
screen "Dev_VD2" 800x480, template "Settings"
   TextField "Text field_10" at 472,32 size 34x18; Text 'ОС.О'
   TextField "Text field_4" at 510,10 size 77x22; Text 'Сигналы:'
   Button "Button_21" at 508,32 size 60x20; TextOff 'Text'; Authorization "User administration"; PictureList "ON_OFF"
      on Click: InvertBit("V_x_Use_Open")
      ProcessValue <- "V_x_Use_Open"
   Button "Button_22" at 508,56 size 60x20; TextOff 'Text'; PictureList "ON_OFF"; Authorization "User administration"
      on Click: InvertBit("V_x_Use_Close")
      ProcessValue <- "V_x_Use_Close"
   Button "Button_27" at 452,31 size 20x20; TextOff 'Text'; Authorization "User administration"; PictureList "signal_green"
      ProcessValue <- "V_x_FB_Open"
   GraphicIOField "Graphic I/O field_5" at 169,56 size 50x50; PictureList "Valve_Hor"
      ProcessValue <- "V_x_Status"
   TextField "Text field_6" at 472,56 size 31x18; Text 'ОС.З'
   Button "Button_12" at 452,55 size 20x20; TextOff 'Text'; Authorization "User administration"; PictureList "signal_green"
      ProcessValue <- "V_x_FB_Close"
   Button "Button_2" at 574,32 size 20x20; TextOff 'Text'; Authorization "User administration"; PictureList "ok_green"
      on Release: InvertBit("V_x_Inv_Open")
      ProcessValue <- "V_x_Inv_Open"
   Button "Button_3" at 574,56 size 20x20; TextOff 'Text'; Authorization "User administration"; PictureList "ok_green"
      on Release: InvertBit("V_x_Inv_Close")
      ProcessValue <- "V_x_Inv_Close"
   IOField "I/O field_1" at 615,30 size 30x24; Authorization "Developer"; FormatPattern 99
      ProcessValue <- "V_x_Indirect_BYTE_FB_Open"
   IOField "I/O field_6" at 655,30 size 20x24; Authorization "Developer"; FormatPattern 9
      ProcessValue <- "V_x_Indirect_BIT_FB_Open"
   TextField "Text field_11" at 601,30 size 13x23; Text 'I'
   TextField "Text field_1" at 644,30 size 13x23; Text '.'
   IOField "I/O field_2" at 615,54 size 30x24; Authorization "Developer"; FormatPattern 99
      ProcessValue <- "V_x_Indirect_BYTE_FB_Close"
   IOField "I/O field_3" at 655,54 size 20x24; Authorization "Developer"; FormatPattern 9
      ProcessValue <- "V_x_Indirect_BIT_FB_Close"
   TextField "Text field_7" at 601,54 size 13x23; Text 'I'
   TextField "Text field_8" at 644,54 size 13x23; Text '.'
   IOField "I/O field_4" at 615,78 size 30x24; Authorization "Developer"; FormatPattern 99
      ProcessValue <- "V_x_Indirect_BYTE_CMD_Open"
   IOField "I/O field_7" at 655,78 size 20x24; Authorization "Developer"; FormatPattern 9
      ProcessValue <- "V_x_Indirect_BIT_CMD_Open"
   TextField "Text field_9" at 599,78 size 17x23; Text 'Q'
   TextField "Text field_13" at 644,78 size 13x23; Text '.'
   TextField "Text field_3" at 472,80 size 65x18; Text 'Открыть / CMD Откр'
   Button "Button_5" at 452,79 size 20x20; TextOff 'Text'; Authorization "User administration"; PictureList "signal_green"
      ProcessValue <- "V_x_CMD_Open"
   IOField "I/O field_8" at 170,11 size 171x26; FormatPattern ????????????????
      ProcessValue <- "Vx_Name"
   Button "Button_14" at 538,142 size 142x20; TextOff 'Фиксация'; Authorization "User administration"; TextList "Air_V"
      on Click: InvertBit("V_x_Use_Electro")
      Appearance <- "V_x_Use_Electro"
      ProcessValue <- "V_x_Use_Electro"
   Button "Button_28" at 540,80 size 60x20; TextOff 'Text'; Authorization "User administration"; PictureList "ON_OFF"
      on Click: InvertBit("V_x_Use_CMD_Open")
      ProcessValue <- "V_x_Use_CMD_Open"
   IOField "I/O field_9" at 615,102 size 30x24; Authorization "Developer"; FormatPattern 99
      ProcessValue <- "V_x_Indirect_BYTE_CMD_Close"
   IOField "I/O field_10" at 655,102 size 20x24; Authorization "Developer"; FormatPattern 9
      ProcessValue <- "V_x_Indirect_BIT_CMD_Close"
   TextField "Text field_12" at 599,102 size 17x23; Text 'Q'
   TextField "Text field_14" at 644,102 size 13x23; Text '.'
   TextField "Text field_16" at 472,104 size 62x18; Text 'Закрыть / CMD Закр'
   Button "Button_20" at 452,103 size 20x20; TextOff 'Text'; Authorization "User administration"; PictureList "signal_green"
      ProcessValue <- "V_x_CMD_Close"
   Button "Button_30" at 539,108 size 60x20; TextOff 'Text'; PictureList "ON_OFF"; Authorization "User administration"
      on Click: InvertBit("V_x_Use_CMD_Close")
      ProcessValue <- "V_x_Use_CMD_Close"
   Button "Button_1" at 165,265 size 112x32; TextOff 'DB 700'; Authorization "User administration"
      on Release: SetTag("Vx", 700); SetTag("Vx_Name", 'DB 700')
      Visibility <- "Support_DB_All_VD2s"
      Appearance <- "Vx"
   Button "Button_4" at 165,305 size 112x32; TextOff 'DB 701'; Authorization "User administration"
      on Release: SetTag("Vx", 701); SetTag("Vx_Name", 'DB 701')
      Visibility <- "Support_DB_All_VD2s"
      Appearance <- "Vx"
   Button "Button_17" at 165,345 size 112x32; TextOff 'DB 702'; Authorization "User administration"
      on Release: SetTag("Vx", 702); SetTag("Vx_Name", 'DB 702')
      Visibility <- "Support_DB_All_VD2s"
      Appearance <- "Vx"
   Button "Button_6" at 165,385 size 112x32; TextOff 'DB 703'; Authorization "User administration"
      on Release: SetTag("Vx", 703); SetTag("Vx_Name", 'DB 703')
      Visibility <- "Support_DB_All_VD2s"
      Appearance <- "Vx"
   Button "Button_15" at 443,265 size 112x32; TextOff 'DB 710'; Authorization "User administration"
      on Release: SetTag("Vx", 710); SetTag("Vx_Name", 'DB 710')
      Visibility <- "Support_DB_All_VD2s"
      Appearance <- "Vx"
   Button "Button_18" at 443,305 size 112x32; TextOff 'DB 711'; Authorization "User administration"
      on Release: SetTag("Vx", 711); SetTag("Vx_Name", 'DB 711')
      Visibility <- "Support_DB_All_VD2s"
      Appearance <- "Vx"
   Button "Button_23" at 443,345 size 112x32; TextOff 'DB 712'; Authorization "User administration"
      on Release: SetTag("Vx", 712); SetTag("Vx_Name", 'DB 712')
      Visibility <- "Support_DB_All_VD2s"
      Appearance <- "Vx"
   Button "Button_24" at 443,385 size 112x32; TextOff 'DB 713'; Authorization "User administration"
      on Release: SetTag("Vx", 713); SetTag("Vx_Name", 'DB 713')
      Visibility <- "Support_DB_All_VD2s"
      Appearance <- "Vx"
   Button "Button_25" at 443,425 size 112x32; TextOff 'DB 714'; Authorization "User administration"
      on Release: SetTag("Vx", 714); SetTag("Vx_Name", 'DB 714')
      Visibility <- "Support_DB_All_VD2s"
      Appearance <- "Vx"
   Button "Button_26" at 583,344 size 112x32; TextOff 'DB 717'; Authorization "User administration"
      on Release: SetTag("Vx", 717); SetTag("Vx_Name", 'DB 717')
      Visibility <- "Support_DB_All_VD2s"
      Appearance <- "Vx"
   Button "Button_29" at 583,384 size 112x32; TextOff 'DB 718'; Authorization "User administration"
      on Release: SetTag("Vx", 718); SetTag("Vx_Name", 'DB 718')
      Visibility <- "Support_DB_All_VD2s"
      Appearance <- "Vx"
   Button "Button_31" at 583,264 size 112x32; TextOff 'DB 715'; Authorization "User administration"
      on Release: SetTag("Vx", 715); SetTag("Vx_Name", 'DB 715')
      Visibility <- "Support_DB_All_VD2s"
      Appearance <- "Vx"
   Button "Button_32" at 583,304 size 112x32; TextOff 'DB 716'; Authorization "User administration"
      on Release: SetTag("Vx", 716); SetTag("Vx_Name", 'DB 716')
      Visibility <- "Support_DB_All_VD2s"
      Appearance <- "Vx"
   Button "Button_33" at 165,425 size 112x32; TextOff 'DB 704'; Authorization "User administration"
      on Release: SetTag("Vx", 704); SetTag("Vx_Name", 'DB 704')
      Visibility <- "Support_DB_All_VD2s"
      Appearance <- "Vx"
   Button "Button_34" at 583,424 size 112x32; TextOff 'DB 719'; Authorization "User administration"
      on Release: SetTag("Vx", 719); SetTag("Vx_Name", 'DB 719')
      Visibility <- "Support_DB_All_VD2s"
      Appearance <- "Vx"
   Button "Button_35" at 304,265 size 112x32; TextOff 'DB 705'; Authorization "User administration"
      on Release: SetTag("Vx", 705); SetTag("Vx_Name", 'DB 705')
      Visibility <- "Support_DB_All_VD2s"
      Appearance <- "Vx"
   Button "Button_36" at 304,305 size 112x32; TextOff 'DB 706'; Authorization "User administration"
      on Release: SetTag("Vx", 706); SetTag("Vx_Name", 'DB 706')
      Visibility <- "Support_DB_All_VD2s"
      Appearance <- "Vx"
   Button "Button_37" at 304,345 size 112x32; TextOff 'DB 707'; Authorization "User administration"
      on Release: SetTag("Vx", 707); SetTag("Vx_Name", 'DB 707')
      Visibility <- "Support_DB_All_VD2s"
      Appearance <- "Vx"
   Button "Button_38" at 304,385 size 112x32; TextOff 'DB 708'; Authorization "User administration"
      on Release: SetTag("Vx", 708); SetTag("Vx_Name", 'DB 708')
      Visibility <- "Support_DB_All_VD2s"
      Appearance <- "Vx"
   Button "Button_39" at 304,425 size 112x32; TextOff 'DB 709'; Authorization "User administration"
      on Release: SetTag("Vx", 709); SetTag("Vx_Name", 'DB 709')
      Visibility <- "Support_DB_All_VD2s"
      Appearance <- "Vx"
   Button "Button_7" at 251,41 size 90x22; TextOff 'Авто'; TextList "Hand"; Authorization "Operate"
      on Click: InvertBit("V_x_CMD_Hand")
      Appearance <- "V_x_CMD_Hand"
      ProcessValue <- "V_x_CMD_Hand"
   Button "Button_8" at 297,66 size 44x40; TextOff 'Закр / Стоп'; Authorization "Operate"
      on Click: ResetBit("V_x_CMD_Start_M")
   Button "Button_13" at 251,66 size 44x40; TextOff 'Откр / Пуск'; Authorization "Operate"
      on Click: SetBit("V_x_CMD_Start_M")
      Appearance <- "V_x_CMD_Start_M"
   TextField "Text field_15" at 348,12 size 99x18; Text 'Ожидание ОС, с'
   GraphicView "Graphic view_1" at 220,42 size 25x25; Picture "z2use_3"
      Visibility <- "V_x_CMD_Hand"
   GraphicView "Graphic view_8" at 220,131 size 25x25; Picture "Force_F"
      Visibility <- "V_x_CMD_Force"
   GraphicView "Graphic view_11" at 220,86 size 25x25; Picture "lock_32x32_1"
      Visibility <- "V_x_CMD_Lock"
   TextField "Text field_2" at 347,34 size 37x18; Text 'Откр. / Старт'
   IOField "I/O field_5" at 386,32 size 30x20; Authorization "User administration"; FormatPattern 99
      ProcessValue <- "V_x_Wait_On_SP"
   IOField "I/O field_12" at 386,55 size 30x20; Authorization "User administration"; FormatPattern 99
      ProcessValue <- "V_x_Wait_Off_SP"
   TextField "Text field_5" at 347,55 size 34x18; Text 'Закр. / Стоп'
   IOField "I/O field_13" at 416,32 size 30x20; FormatPattern 99
      ProcessValue <- "V_x_Wait_On_Now"
   IOField "I/O field_14" at 416,55 size 30x20; FormatPattern 99
      ProcessValue <- "V_x_Wait_Off_Now"
   Button "Button_11" at 251,109 size 90x20; TextOff 'Принудит.'; Authorization "User administration"
      on Click: InvertBit("V_x_CMD_Force")
      Appearance <- "V_x_CMD_Force"
   GraphicView "Graphic view_55" at 169,134 size 24x21; Picture "local"
      Visibility <- "V_x_CMD_Local"
   Button "Button_19" at 251,132 size 90x22; TextOff 'Сброс аварий'; Authorization "Operate"
      on Click: SetBit("V_x_CMD_Reset")
   GraphicView "Graphic view_3" at 194,131 size 25x25; Picture "service"
      Visibility <- "V_x_CMD_Service"
   TextField "Text field_17" at 348,84 size 74x18; Text 'Задержка, с'
   TextField "Text field_18" at 347,106 size 37x18; Text 'Откр. / Пуск'
   IOField "I/O field_11" at 386,104 size 30x20; Authorization "User administration"; FormatPattern 99
      ProcessValue <- "V_x_Delay_On_SP"
   IOField "I/O field_16" at 386,127 size 30x20; Authorization "User administration"; FormatPattern 99
      ProcessValue <- "V_x_Delay_Off_SP"
   TextField "Text field_20" at 347,127 size 34x18; Text 'Закр. / Стоп'
   IOField "I/O field_17" at 416,104 size 30x20; FormatPattern 99
      ProcessValue <- "V_x_Delay_On_Now"
   IOField "I/O field_18" at 416,127 size 30x20; FormatPattern 99
      ProcessValue <- "V_x_Delay_Off_Now"
   TextField "Text field_19" at 454,144 size 82x18; Text 'Тип привода:'
   SymbolicIOField "Symbolic I/O field_1" at 113,464 size 75x16; TextOn '1'; TextOff '0'; TextList "Hand"
      ProcessValue <- "V_x_CMD_Hand"
   TextField "Text field_21" at 211,464 size 75x16; Text 'Открыть'
      Visibility <- "V_x_CMD_Hand"
   TextField "Text field_22" at 311,464 size 75x16; Text 'Закрыть'
      Visibility <- "V_x_CMD_Hand"
   TextField "Text field_23" at 610,464 size 75x16; Text 'Сброс аварий'
   Softkey "Softkey_F2" at 0,0 size 0x0
      on KeyDown: InvertBit("V_x_CMD_Hand")
   Softkey "Softkey_F3" at 0,0 size 0x0
      on KeyDown: SetBit("V_x_CMD_Start_M")
   Softkey "Softkey_F4" at 0,0 size 0x0
      on KeyDown: ResetBit("V_x_CMD_Start_M")
   Softkey "Softkey_F7" at 0,0 size 0x0
      on KeyDown: SetBit("V_x_CMD_Reset")

screen "Dev_MDA" 800x480, template "Settings"
   Rectangle "Rectangle_1" at 165,7 size 520x253
      Appearance <- "M_x_CMD_Sim"
   IOField "I/O field_17" at 168,226 size 80x30; Authorization "User administration"; FormatPattern s999.99
      Appearance <- "M_x_CMD_Hand"
      ProcessValue <- "MA_x_SP_M"
   TextField "Text field_19" at 181,208 size 48x18; Text 'Уставка'
   TextField "Text field_38" at 358,216 size 75x18; Text 'Тип выхода:'
      Visibility <- "AI_x_Use_RTD"
   IOField "I/O field_32" at 347,236 size 42x20; Authorization "User administration"; FormatPattern 99.99
      Visibility <- "AI_x_Use_RTD"
      ProcessValue <- "MA_x_VmA"
   Button "Button_10" at 393,236 size 56x20; TextOff 'Авто'; Authorization "Developer"; TextList "VmA_2"
      on Click: function_dd21b452("MA_x_Output_Type", 1)
      Visibility <- "AI_x_Use_RTD"
      ProcessValue <- "MA_x_Output_Type"
   TextField "Text field_20" at 525,102 size 107x18; Text 'Масштабирование'
   TextField "Text field_21" at 560,114 size 18x18; Text 'от'
   IOField "I/O field_19" at 541,132 size 57x20; Authorization "User administration"; FormatPattern s999.99
      ProcessValue <- "MA_x_Converter_Min_In"
   TextField "Text field_22" at 613,114 size 19x18; Text 'до'
   IOField "I/O field_20" at 602,132 size 57x20; Authorization "User administration"; FormatPattern s999.99
      ProcessValue <- "MA_x_Converter_Max_In"
   TextField "Text field_28" at 489,133 size 52x18; Text 'Уставка:'
   IOField "I/O field_23" at 541,156 size 57x20; Authorization "User administration"; FormatPattern 99999
      ProcessValue <- "MA_x_Converter_Min_Out"
   IOField "I/O field_26" at 602,156 size 57x20; Authorization "User administration"; FormatPattern 99999
      ProcessValue <- "MA_x_Converter_Max_Out"
   TextField "Text field_29" at 499,157 size 32x18; Text 'ПЛК:'
   IOField "I/O field_27" at 482,235 size 57x20; Authorization "Developer"; FormatPattern 999
      ProcessValue <- "MA_x_Indirect_BYTE_SP"
   TextField "Text field_36" at 456,236 size 26x18; Text 'QW'
   GraphicIOField "Graphic I/O field_2" at 172,43 size 43x85; PictureList "Motor"
      ProcessValue <- "M_x_Status"
   Button "Button_7" at 251,41 size 90x22; TextOff 'Авто'; TextList "Hand"; Authorization "Operate"
      on Click: InvertBit("M_x_CMD_Hand")
      Appearance <- "M_x_CMD_Hand"
      ProcessValue <- "M_x_CMD_Hand"
   Button "Button_8" at 297,66 size 44x40; TextOff 'Стоп'; Authorization "Operate"
      on Click: ResetBit("M_x_CMD_Start_M")
   Button "Button_13" at 251,66 size 44x40; TextOff 'Пуск'; Authorization "Operate"
      on Click: SetBit("M_x_CMD_Start_M")
      Appearance <- "M_x_CMD_Start_M"
   TextField "Text field_15" at 348,12 size 99x18; Text 'Ожидание ОС, с'
   GraphicView "Graphic view_1" at 220,42 size 25x25; Picture "z2use_3"
      Visibility <- "M_x_CMD_Hand"
   GraphicView "Graphic view_8" at 220,131 size 25x25; Picture "Force_F"
      Visibility <- "M_x_CMD_Force"
   GraphicView "Graphic view_11" at 220,86 size 25x25; Picture "lock_32x32_1"
      Visibility <- "M_x_CMD_Lock"
   TextField "Text field_3" at 474,31 size 20x18; Text 'QF'
   TextField "Text field_10" at 474,56 size 21x18; Text 'KM'
   TextField "Text field_12" at 474,82 size 29x18; Text 'CMD'
   TextField "Text field_4" at 478,10 size 197x22; Text 'Конфигурация сигналов:'
   Button "Button_21" at 508,32 size 60x20; TextOff 'Text'; PictureList "ON_OFF"; Authorization "User administration"
      on Click: InvertBit("M_x_Use_QF")
      ProcessValue <- "M_x_Use_QF"
   Button "Button_22" at 508,56 size 60x20; TextOff 'Text'; Authorization "User administration"; PictureList "ON_OFF"
      on Click: InvertBit("M_x_Use_KM")
      ProcessValue <- "M_x_Use_KM"
   Button "Button_26" at 454,31 size 20x20; TextOff 'Text'; Authorization "User administration"; PictureList "signal_green"
      ProcessValue <- "M_x_FB_QF"
   Button "Button_27" at 454,55 size 20x20; TextOff 'Text'; Authorization "User administration"; PictureList "signal_green"
      ProcessValue <- "M_x_FB_KM"
   Button "Button_29" at 454,80 size 20x20; TextOff 'Text'; Authorization "User administration"; PictureList "signal_green"
      ProcessValue <- "M_x_CMD"
   TextField "Text field_2" at 347,34 size 37x18; Text 'Старт'
   IOField "I/O field_5" at 386,32 size 30x20; Authorization "User administration"; FormatPattern 99
      ProcessValue <- "M_x_Wait_On_SP"
   IOField "I/O field_12" at 386,55 size 30x20; Authorization "User administration"; FormatPattern 99
      ProcessValue <- "M_x_Wait_Off_SP"
   TextField "Text field_5" at 347,55 size 32x18; Text 'Стоп'
   IOField "I/O field_13" at 416,32 size 30x20; FormatPattern 99
      ProcessValue <- "M_x_Wait_On_Now"
   IOField "I/O field_14" at 416,55 size 30x20; FormatPattern 99
      ProcessValue <- "M_x_Wait_Off_Now"
   Button "Button_11" at 251,109 size 90x20; TextOff 'Принудит.'; Authorization "User administration"
      on Click: InvertBit("M_x_CMD_Force")
      Appearance <- "M_x_CMD_Force"
   Button "Button_2" at 574,31 size 20x20; TextOff 'Text'; Authorization "User administration"; PictureList "ok_green"
      on Click: InvertBit("M_x_Inv_QF")
      ProcessValue <- "M_x_Inv_QF"
   Button "Button_3" at 574,55 size 20x20; TextOff 'Text'; PictureList "ok_green"; Authorization "User administration"
      on Click: InvertBit("M_x_Inv_KM")
      ProcessValue <- "M_x_Inv_KM"
   IOField "I/O field_1" at 615,30 size 30x24; Authorization "Developer"; FormatPattern 99
      ProcessValue <- "M_x_Indirect_BYTE_FB_QF"
   IOField "I/O field_6" at 655,30 size 22x24; Authorization "Developer"; FormatPattern 9
      ProcessValue <- "M_x_Indirect_BIT_FB_QF"
   TextField "Text field_11" at 599,30 size 13x23; Text 'I'
   TextField "Text field_6" at 644,30 size 13x23; Text '.'
   IOField "I/O field_2" at 615,54 size 30x24; Authorization "Developer"; FormatPattern 99
      ProcessValue <- "M_x_Indirect_BYTE_FB_KM"
   IOField "I/O field_3" at 655,54 size 22x24; Authorization "Developer"; FormatPattern 9
      ProcessValue <- "M_x_Indirect_BIT_FB_KM"
   TextField "Text field_7" at 599,54 size 13x23; Text 'I'
   TextField "Text field_8" at 644,54 size 13x23; Text '.'
   IOField "I/O field_4" at 615,78 size 30x24; Authorization "Developer"; FormatPattern 99
      ProcessValue <- "M_x_Indirect_BYTE_CMD"
   IOField "I/O field_7" at 655,78 size 22x24; Authorization "Developer"; FormatPattern 9
      ProcessValue <- "M_x_Indirect_BIT_CMD"
   TextField "Text field_9" at 597,78 size 17x23; Text 'Q'
   TextField "Text field_13" at 644,78 size 13x23; Text '.'
   IOField "I/O field_8" at 170,11 size 171x26; FormatPattern ????????????????
      ProcessValue <- "Mx_Name"
   Button "Button_4" at 508,80 size 60x20; TextOff 'Text'; Authorization "User administration"; PictureList "ON_OFF"
      on Click: InvertBit("M_x_Indirect_CMD")
      ProcessValue <- "M_x_Indirect_CMD"
   TextField "Text field_14" at 168,158 size 79x18; Text 'Наработка, ч'
   IOField "I/O field_9" at 251,158 size 90x20; FormatPattern 9999999999
      ProcessValue <- "M_x_OpTime_All_h"
   TextField "Text field_18" at 170,183 size 108x18; Text 'Сервис каждые, ч'
   IOField "I/O field_15" at 293,181 size 48x22; FormatPattern 99999
      ProcessValue <- "M_x_OpTime_SP_h"
   Button "Button_16" at 410,181 size 82x22; TextOff 'Сервис'; Authorization "Operate"
      on Click: SetBit("M_x_CMD_ResetOpTime")
      Appearance <- "M_x_OpTime_Alarm"
   TextField "Text field_1" at 494,183 size 122x18; Text 'Контроль наработки'
   Button "Button_18" at 617,182 size 60x20; TextOff 'Text'; PictureList "ON_OFF"; Authorization "User administration"
      on Click: InvertBit("M_x_Use_OpTime")
      ProcessValue <- "M_x_Use_OpTime"
   IOField "I/O field_10" at 357,181 size 48x22; FormatPattern 99999
      ProcessValue <- "M_x_OpTime_Now_h"
   TextField "Text field_16" at 344,183 size 10x18; Text '/'
   GraphicView "Graphic view_55" at 169,134 size 24x21; Picture "local"
      Visibility <- "M_x_CMD_Local"
   Button "Button_9" at 251,132 size 90x22; TextOff 'Сброс аварий'; TextList "Hand_1"; Authorization "Operate"
      on Click: SetBit("M_x_CMD_Reset")
      ProcessValue <- "MA_x_CMD_Hand"
   GraphicView "Graphic view_3" at 194,131 size 25x25; Picture "service"
      Visibility <- "M_x_CMD_Service"
   TextField "Text field_17" at 348,84 size 74x18; Text 'Задержка, с'
   TextField "Text field_23" at 347,106 size 31x18; Text 'Пуск'
   IOField "I/O field_11" at 386,104 size 30x20; Authorization "User administration"; FormatPattern 99
      ProcessValue <- "M_x_Delay_On_SP"
   IOField "I/O field_16" at 386,127 size 30x20; Authorization "User administration"; FormatPattern 99
      ProcessValue <- "M_x_Delay_Off_SP"
   TextField "Text field_24" at 347,127 size 32x18; Text 'Стоп'
   IOField "I/O field_18" at 416,104 size 30x20; FormatPattern 99
      ProcessValue <- "M_x_Delay_On_Now"
   IOField "I/O field_21" at 416,127 size 30x20; FormatPattern 99
      ProcessValue <- "M_x_Delay_Off_Now"
   TextField "Text field_25" at 259,208 size 81x18; Text 'Размерность:'
   Button "Button_19" at 258,226 size 80x30; TextOff 'Авто'; TextList "Input_Type"; Authorization "Developer"
      on Click: function_dd21b452("AO_x_Type", 1)
      ProcessValue <- "MA_x_Type"
   Button "Button_1" at 165,265 size 112x32; TextOff 'DB 600'; Authorization "User administration"
      on Release: SetTag("Mx", 600); SetTag("Mx_Name", 'DB 600')
      Visibility <- "Support_DB_All_MDAs"
      Appearance <- "Mx"
   Button "Button_5" at 165,305 size 112x32; TextOff 'DB 601'; Authorization "User administration"
      on Release: SetTag("Mx", 601); SetTag("Mx_Name", 'DB 601')
      Visibility <- "Support_DB_All_MDAs"
      Appearance <- "Mx"
   Button "Button_17" at 165,345 size 112x32; TextOff 'DB 602'; Authorization "User administration"
      on Release: SetTag("Mx", 602); SetTag("Mx_Name", 'DB 602')
      Visibility <- "Support_DB_All_MDAs"
      Appearance <- "Mx"
   Button "Button_6" at 165,385 size 112x32; TextOff 'DB 603'; Authorization "User administration"
      on Release: SetTag("Mx", 603); SetTag("Mx_Name", 'DB 603')
      Visibility <- "Support_DB_All_MDAs"
      Appearance <- "Mx"
   Button "Button_12" at 443,265 size 112x32; TextOff 'DB 610'; Authorization "User administration"
      on Release: SetTag("Mx", 610); SetTag("Mx_Name", 'DB 610')
      Visibility <- "Support_DB_All_MDAs"
      Appearance <- "Mx"
   Button "Button_14" at 443,305 size 112x32; TextOff 'DB 611'; Authorization "User administration"
      on Release: SetTag("Mx", 611); SetTag("Mx_Name", 'DB 611')
      Visibility <- "Support_DB_All_MDAs"
      Appearance <- "Mx"
   Button "Button_15" at 443,345 size 112x32; TextOff 'DB 612'; Authorization "User administration"
      on Release: SetTag("Mx", 612); SetTag("Mx_Name", 'DB 612')
      Visibility <- "Support_DB_All_MDAs"
      Appearance <- "Mx"
   Button "Button_20" at 443,385 size 112x32; TextOff 'DB 613'; Authorization "User administration"
      on Release: SetTag("Mx", 613); SetTag("Mx_Name", 'DB 613')
      Visibility <- "Support_DB_All_MDAs"
      Appearance <- "Mx"
   Button "Button_23" at 443,425 size 112x32; TextOff 'DB 614'; Authorization "User administration"
      on Release: SetTag("Mx", 614); SetTag("Mx_Name", 'DB 614')
      Visibility <- "Support_DB_All_MDAs"
      Appearance <- "Mx"
   Button "Button_24" at 583,344 size 112x32; TextOff 'DB 617'; Authorization "User administration"
      on Release: SetTag("Mx", 617); SetTag("Mx_Name", 'DB 617')
      Visibility <- "Support_DB_All_MDAs"
      Appearance <- "Mx"
   Button "Button_25" at 583,384 size 112x32; TextOff 'DB 618'; Authorization "User administration"
      on Release: SetTag("Mx", 618); SetTag("Mx_Name", 'DB 618')
      Visibility <- "Support_DB_All_MDAs"
      Appearance <- "Mx"
   Button "Button_28" at 583,264 size 112x32; TextOff 'DB 615'; Authorization "User administration"
      on Release: SetTag("Mx", 615); SetTag("Mx_Name", 'DB 615')
      Visibility <- "Support_DB_All_MDAs"
      Appearance <- "Mx"
   Button "Button_30" at 583,304 size 112x32; TextOff 'DB 616'; Authorization "User administration"
      on Release: SetTag("Mx", 616); SetTag("Mx_Name", 'DB 616')
      Visibility <- "Support_DB_All_MDAs"
      Appearance <- "Mx"
   Button "Button_31" at 165,425 size 112x32; TextOff 'DB 604'; Authorization "User administration"
      on Release: SetTag("Mx", 604); SetTag("Mx_Name", 'DB 604')
      Visibility <- "Support_DB_All_MDAs"
      Appearance <- "Mx"
   Button "Button_32" at 583,424 size 112x32; TextOff 'DB 619'; Authorization "User administration"
      on Release: SetTag("Mx", 619); SetTag("Mx_Name", 'DB 619')
      Visibility <- "Support_DB_All_MDAs"
      Appearance <- "Mx"
   Button "Button_33" at 304,265 size 112x32; TextOff 'DB 605'; Authorization "User administration"
      on Release: SetTag("Mx", 605); SetTag("Mx_Name", 'DB 605')
      Visibility <- "Support_DB_All_MDAs"
      Appearance <- "Mx"
   Button "Button_34" at 304,305 size 112x32; TextOff 'DB 606'; Authorization "User administration"
      on Release: SetTag("Mx", 606); SetTag("Mx_Name", 'DB 606')
      Visibility <- "Support_DB_All_MDAs"
      Appearance <- "Mx"
   Button "Button_35" at 304,345 size 112x32; TextOff 'DB 607'; Authorization "User administration"
      on Release: SetTag("Mx", 607); SetTag("Mx_Name", 'DB 607')
      Visibility <- "Support_DB_All_MDAs"
      Appearance <- "Mx"
   Button "Button_36" at 304,385 size 112x32; TextOff 'DB 608'; Authorization "User administration"
      on Release: SetTag("Mx", 608); SetTag("Mx_Name", 'DB 608')
      Visibility <- "Support_DB_All_MDAs"
      Appearance <- "Mx"
   Button "Button_37" at 304,425 size 112x32; TextOff 'DB 609'; Authorization "User administration"
      on Release: SetTag("Mx", 609); SetTag("Mx_Name", 'DB 609')
      Visibility <- "Support_DB_All_MDAs"
      Appearance <- "Mx"
   SymbolicIOField "Symbolic I/O field_1" at 113,464 size 75x16; TextOn '1'; TextOff '0'; TextList "Hand"
      ProcessValue <- "M_x_CMD_Hand"
   TextField "Text field_26" at 211,464 size 75x16; Text 'Пуск'
      Visibility <- "M_x_CMD_Hand"
   TextField "Text field_27" at 311,464 size 75x16; Text 'Стоп'
      Visibility <- "M_x_CMD_Hand"
   TextField "Text field_30" at 610,464 size 75x16; Text 'Сброс аварий'
   Softkey "Softkey_F2" at 0,0 size 0x0
      on KeyDown: InvertBit("M_x_CMD_Hand")
   Softkey "Softkey_F3" at 0,0 size 0x0
      on KeyDown: SetBit("M_x_CMD_Start_M")
   Softkey "Softkey_F4" at 0,0 size 0x0
      on KeyDown: ResetBit("M_x_CMD_Start_M")
   Softkey "Softkey_F7" at 0,0 size 0x0
      on KeyDown: SetBit("M_x_CMD_Reset")

screen "Dev_MD" 800x480, template "Settings"
   Rectangle "Rectangle_1" at 165,7 size 520x200
      Appearance <- "M_x_CMD_Sim"
   GraphicIOField "Graphic I/O field_2" at 172,43 size 43x85; PictureList "Motor"
      ProcessValue <- "M_x_Status"
   Button "Button_7" at 251,41 size 90x22; TextOff 'Авто'; Authorization "Operate"; TextList "Hand"
      on Click: InvertBit("M_x_CMD_Hand")
      Appearance <- "M_x_CMD_Hand"
      ProcessValue <- "M_x_CMD_Hand"
   Button "Button_8" at 297,66 size 44x40; TextOff 'Стоп'; Authorization "Operate"
      on Click: ResetBit("M_x_CMD_Start_M")
   Button "Button_13" at 251,66 size 44x40; TextOff 'Пуск'; Authorization "Operate"
      on Click: SetBit("M_x_CMD_Start_M")
      Appearance <- "M_x_CMD_Start_M"
   TextField "Text field_15" at 348,12 size 99x18; Text 'Ожидание ОС, с'
   GraphicView "Graphic view_1" at 220,42 size 25x25; Picture "z2use_3"
      Visibility <- "M_x_CMD_Hand"
   GraphicView "Graphic view_8" at 220,131 size 25x25; Picture "Force_F"
      Visibility <- "M_x_CMD_Force"
   GraphicView "Graphic view_11" at 220,86 size 25x25; Picture "lock_32x32_1"
      Visibility <- "M_x_CMD_Lock"
   TextField "Text field_3" at 474,31 size 20x18; Text 'QF'
   TextField "Text field_10" at 474,56 size 21x18; Text 'KM'
   TextField "Text field_12" at 474,82 size 29x18; Text 'CMD'
   TextField "Text field_4" at 478,10 size 197x22; Text 'Конфигурация сигналов:'
   Button "Button_21" at 508,32 size 60x20; TextOff 'Text'; Authorization "User administration"; PictureList "ON_OFF"
      on Click: InvertBit("M_x_Use_QF")
      ProcessValue <- "M_x_Use_QF"
   Button "Button_22" at 508,56 size 60x20; TextOff 'Text'; PictureList "ON_OFF"; Authorization "User administration"
      on Click: InvertBit("M_x_Use_KM")
      ProcessValue <- "M_x_Use_KM"
   Button "Button_26" at 454,31 size 20x20; TextOff 'Text'; Authorization "User administration"; PictureList "signal_green"
      ProcessValue <- "M_x_FB_QF"
   Button "Button_27" at 454,55 size 20x20; TextOff 'Text'; Authorization "User administration"; PictureList "signal_green"
      ProcessValue <- "M_x_FB_KM"
   Button "Button_29" at 454,80 size 20x20; TextOff 'Text'; Authorization "User administration"; PictureList "signal_green"
      ProcessValue <- "M_x_CMD"
   TextField "Text field_2" at 347,34 size 37x18; Text 'Старт'
   IOField "I/O field_5" at 386,32 size 30x20; Authorization "User administration"; FormatPattern 99
      ProcessValue <- "M_x_Wait_On_SP"
   IOField "I/O field_12" at 386,55 size 30x20; Authorization "User administration"; FormatPattern 99
      ProcessValue <- "M_x_Wait_Off_SP"
   TextField "Text field_5" at 347,55 size 32x18; Text 'Стоп'
   IOField "I/O field_13" at 416,32 size 30x20; FormatPattern 99
      ProcessValue <- "M_x_Wait_On_Now"
   IOField "I/O field_14" at 416,55 size 30x20; FormatPattern 99
      ProcessValue <- "M_x_Wait_Off_Now"
   Button "Button_11" at 251,109 size 90x20; TextOff 'Принудит.'; Authorization "User administration"
      on Click: InvertBit("M_x_CMD_Force")
      Appearance <- "M_x_CMD_Force"
   Button "Button_2" at 574,31 size 20x20; TextOff 'Text'; Authorization "User administration"; PictureList "ok_green"
      on Click: InvertBit("M_x_Inv_QF")
      ProcessValue <- "M_x_Inv_QF"
   Button "Button_3" at 574,55 size 20x20; TextOff 'Text'; Authorization "User administration"; PictureList "ok_green"
      on Click: InvertBit("M_x_Inv_KM")
      ProcessValue <- "M_x_Inv_KM"
   IOField "I/O field_1" at 615,30 size 30x24; Authorization "Developer"; FormatPattern 99
      ProcessValue <- "M_x_Indirect_BYTE_FB_QF"
   IOField "I/O field_6" at 655,30 size 22x24; Authorization "Developer"; FormatPattern 9
      ProcessValue <- "M_x_Indirect_BIT_FB_QF"
   TextField "Text field_11" at 599,30 size 13x23; Text 'I'
   TextField "Text field_6" at 644,30 size 13x23; Text '.'
   IOField "I/O field_2" at 615,54 size 30x24; Authorization "Developer"; FormatPattern 99
      ProcessValue <- "M_x_Indirect_BYTE_FB_KM"
   IOField "I/O field_3" at 655,54 size 22x24; Authorization "Developer"; FormatPattern 9
      ProcessValue <- "M_x_Indirect_BIT_FB_KM"
   TextField "Text field_7" at 599,54 size 13x23; Text 'I'
   TextField "Text field_8" at 644,54 size 13x23; Text '.'
   IOField "I/O field_4" at 615,78 size 30x24; Authorization "Developer"; FormatPattern 99
      ProcessValue <- "M_x_Indirect_BYTE_CMD"
   IOField "I/O field_7" at 655,78 size 22x24; Authorization "Developer"; FormatPattern 9
      ProcessValue <- "M_x_Indirect_BIT_CMD"
   TextField "Text field_9" at 597,78 size 17x23; Text 'Q'
   TextField "Text field_13" at 644,78 size 13x23; Text '.'
   IOField "I/O field_8" at 170,11 size 171x26; FormatPattern ????????????????
      ProcessValue <- "Mx_Name"
   Button "Button_15" at 508,80 size 60x20; TextOff 'Text'; PictureList "ON_OFF"; Authorization "User administration"
      on Click: InvertBit("M_x_Indirect_CMD")
      ProcessValue <- "M_x_Indirect_CMD"
   TextField "Text field_14" at 168,158 size 79x18; Text 'Наработка, ч'
   IOField "I/O field_9" at 251,158 size 90x20; FormatPattern 9999999999
      ProcessValue <- "M_x_OpTime_All_h"
   TextField "Text field_18" at 170,183 size 108x18; Text 'Сервис каждые, ч'
   IOField "I/O field_15" at 293,181 size 48x22; FormatPattern 99999
      ProcessValue <- "M_x_OpTime_SP_h"
   Button "Button_16" at 410,181 size 82x22; TextOff 'Сервис'; Authorization "Operate"
      on Click: SetBit("M_x_CMD_ResetOpTime")
      Appearance <- "M_x_OpTime_Alarm"
   TextField "Text field_19" at 494,183 size 122x18; Text 'Контроль наработки'
   Button "Button_18" at 617,182 size 60x20; TextOff 'Text'; Authorization "User administration"; PictureList "ON_OFF"
      on Click: InvertBit("M_x_Use_OpTime")
      ProcessValue <- "M_x_Use_OpTime"
   IOField "I/O field_10" at 357,181 size 48x22; FormatPattern 99999
      ProcessValue <- "M_x_OpTime_Now_h"
   TextField "Text field_1" at 344,183 size 10x18; Text '/'
   GraphicView "Graphic view_55" at 169,134 size 24x21; Picture "local"
      Visibility <- "M_x_CMD_Local"
   Button "Button_9" at 251,132 size 90x22; TextOff 'Сброс аварий'; Authorization "Operate"
      on Click: SetBit("M_x_CMD_Reset")
   GraphicView "Graphic view_3" at 194,131 size 25x25; Picture "service"
      Visibility <- "M_x_CMD_Service"
   TextField "Text field_16" at 348,84 size 74x18; Text 'Задержка, с'
   TextField "Text field_17" at 347,106 size 31x18; Text 'Пуск'
   IOField "I/O field_11" at 386,104 size 30x20; Authorization "User administration"; FormatPattern 99
      ProcessValue <- "M_x_Delay_On_SP"
   IOField "I/O field_16" at 386,127 size 30x20; Authorization "User administration"; FormatPattern 99
      ProcessValue <- "M_x_Delay_Off_SP"
   TextField "Text field_20" at 347,127 size 32x18; Text 'Стоп'
   IOField "I/O field_17" at 416,104 size 30x20; FormatPattern 99
      ProcessValue <- "M_x_Delay_On_Now"
   IOField "I/O field_18" at 416,127 size 30x20; FormatPattern 99
      ProcessValue <- "M_x_Delay_Off_Now"
   Button "Button_1" at 165,265 size 112x32; TextOff 'DB 500'; Authorization "User administration"
      on Release: SetTag("Mx", 500); SetTag("Mx_Name", 'DB 500')
      Visibility <- "Support_DB_All_MDs"
      Appearance <- "Mx"
   Button "Button_4" at 165,305 size 112x32; TextOff 'DB 501'; Authorization "User administration"
      on Release: SetTag("Mx", 501); SetTag("Mx_Name", 'DB 501')
      Visibility <- "Support_DB_All_MDs"
      Appearance <- "Mx"
   Button "Button_17" at 165,345 size 112x32; TextOff 'DB 502'; Authorization "User administration"
      on Release: SetTag("Mx", 502); SetTag("Mx_Name", 'DB 502')
      Visibility <- "Support_DB_All_MDs"
      Appearance <- "Mx"
   Button "Button_5" at 165,385 size 112x32; TextOff 'DB 503'; Authorization "User administration"
      on Release: SetTag("Mx", 503); SetTag("Mx_Name", 'DB 503')
      Visibility <- "Support_DB_All_MDs"
      Appearance <- "Mx"
   Button "Button_6" at 443,265 size 112x32; TextOff 'DB 510'; Authorization "User administration"
      on Release: SetTag("Mx", 510); SetTag("Mx_Name", 'DB 510')
      Visibility <- "Support_DB_All_MDs"
      Appearance <- "Mx"
   Button "Button_10" at 443,305 size 112x32; TextOff 'DB 511'; Authorization "User administration"
      on Release: SetTag("Mx", 511); SetTag("Mx_Name", 'DB 511')
      Visibility <- "Support_DB_All_MDs"
      Appearance <- "Mx"
   Button "Button_12" at 443,345 size 112x32; TextOff 'DB 512'; Authorization "User administration"
      on Release: SetTag("Mx", 512); SetTag("Mx_Name", 'DB 512')
      Visibility <- "Support_DB_All_MDs"
      Appearance <- "Mx"
   Button "Button_14" at 443,385 size 112x32; TextOff 'DB 513'; Authorization "User administration"
      on Release: SetTag("Mx", 513); SetTag("Mx_Name", 'DB 513')
      Visibility <- "Support_DB_All_MDs"
      Appearance <- "Mx"
   Button "Button_19" at 443,425 size 112x32; TextOff 'DB 514'; Authorization "User administration"
      on Release: SetTag("Mx", 514); SetTag("Mx_Name", 'DB 514')
      Visibility <- "Support_DB_All_MDs"
      Appearance <- "Mx"
   Button "Button_20" at 583,344 size 112x32; TextOff 'DB 517'; Authorization "User administration"
      on Release: SetTag("Mx", 517); SetTag("Mx_Name", 'DB 517')
      Visibility <- "Support_DB_All_MDs"
      Appearance <- "Mx"
   Button "Button_23" at 583,384 size 112x32; TextOff 'DB 518'; Authorization "User administration"
      on Release: SetTag("Mx", 518); SetTag("Mx_Name", 'DB 518')
      Visibility <- "Support_DB_All_MDs"
      Appearance <- "Mx"
   Button "Button_24" at 583,264 size 112x32; TextOff 'DB 515'; Authorization "User administration"
      on Release: SetTag("Mx", 515); SetTag("Mx_Name", 'DB 515')
      Visibility <- "Support_DB_All_MDs"
      Appearance <- "Mx"
   Button "Button_25" at 583,304 size 112x32; TextOff 'DB 516'; Authorization "User administration"
      on Release: SetTag("Mx", 516); SetTag("Mx_Name", 'DB 516')
      Visibility <- "Support_DB_All_MDs"
      Appearance <- "Mx"
   Button "Button_28" at 165,425 size 112x32; TextOff 'DB 504'; Authorization "User administration"
      on Release: SetTag("Mx", 504); SetTag("Mx_Name", 'DB 504')
      Visibility <- "Support_DB_All_MDs"
      Appearance <- "Mx"
   Button "Button_30" at 583,424 size 112x32; TextOff 'DB 519'; Authorization "User administration"
      on Release: SetTag("Mx", 519); SetTag("Mx_Name", 'DB 519')
      Visibility <- "Support_DB_All_MDs"
      Appearance <- "Mx"
   Button "Button_31" at 304,265 size 112x32; TextOff 'DB 505'; Authorization "User administration"
      on Release: SetTag("Mx", 505); SetTag("Mx_Name", 'DB 505')
      Visibility <- "Support_DB_All_MDs"
      Appearance <- "Mx"
   Button "Button_32" at 304,305 size 112x32; TextOff 'DB 506'; Authorization "User administration"
      on Release: SetTag("Mx", 506); SetTag("Mx_Name", 'DB 506')
      Visibility <- "Support_DB_All_MDs"
      Appearance <- "Mx"
   Button "Button_33" at 304,345 size 112x32; TextOff 'DB 507'; Authorization "User administration"
      on Release: SetTag("Mx", 507); SetTag("Mx_Name", 'DB 507')
      Visibility <- "Support_DB_All_MDs"
      Appearance <- "Mx"
   Button "Button_34" at 304,385 size 112x32; TextOff 'DB 508'; Authorization "User administration"
      on Release: SetTag("Mx", 508); SetTag("Mx_Name", 'DB 508')
      Visibility <- "Support_DB_All_MDs"
      Appearance <- "Mx"
   Button "Button_35" at 304,425 size 112x32; TextOff 'DB 509'; Authorization "User administration"
      on Release: SetTag("Mx", 509); SetTag("Mx_Name", 'DB 509')
      Visibility <- "Support_DB_All_MDs"
      Appearance <- "Mx"
   SymbolicIOField "Symbolic I/O field_1" at 113,464 size 75x16; TextOff '0'; TextOn '1'; TextList "Hand"
      ProcessValue <- "M_x_CMD_Hand"
   TextField "Text field_21" at 211,464 size 75x16; Text 'Пуск'
      Visibility <- "M_x_CMD_Hand"
   TextField "Text field_22" at 311,464 size 75x16; Text 'Стоп'
      Visibility <- "M_x_CMD_Hand"
   TextField "Text field_23" at 610,464 size 75x16; Text 'Сброс аварий'
   Softkey "Softkey_F2" at 0,0 size 0x0
      on KeyDown: InvertBit("M_x_CMD_Hand")
   Softkey "Softkey_F3" at 0,0 size 0x0
      on KeyDown: SetBit("M_x_CMD_Start_M")
   Softkey "Softkey_F4" at 0,0 size 0x0
      on KeyDown: ResetBit("M_x_CMD_Start_M")
   Softkey "Softkey_F7" at 0,0 size 0x0
      on KeyDown: SetBit("M_x_CMD_Reset")

screen "Different jobs" 800x480, template "Main"
   Button "Online" at 36,95 size 159x47; TextOn 'Online'; TextOff 'Online'
      on Release: function_bb44b551(0)
   Button "Offline" at 36,154 size 159x47; TextOn 'Offline'; TextOff 'Offline'
      on Release: function_bb44b551(1)
   Button "Transfer" at 36,213 size 159x47; TextOn 'Transfer'; TextOff 'Transfer'
      on Release: function_bb44b551(2)
   Button "Toggle language" at 36,272 size 159x47; TextOn 'Toggle language'; TextOff 'Toggle language'
      on Release: function_fb9197e8(-1)
   Button "Stop Runtime" at 36,331 size 159x47; TextOn 'Stop Runtime'; TextOff 'Stop Runtime'
      on Release: StopRuntime(0)
   Button "Back" at 1,1 size 159x47; TextOn 'Back'; TextOff 'Back'
      on Release: ActivateScreen("System screens", 0)
   DateTimeField "Date/time field_1" at 448,259 size 111x32
   DateTimeField "Date/time field_2" at 320,259 size 116x32
   TextField "Text field_6" at 560,264 size 18x23; Text 'г.'
   TextField "Text field_2" at 321,232 size 242x23; Text 'Настройка времени панели:'
   DateTimeField "Date/time field_3" at 448,355 size 111x32
      ProcessValue <- "Time_SYS_DB_RD_Time"
   DateTimeField "Date/time field_4" at 320,355 size 116x32
      ProcessValue <- "Time_SYS_DB_RD_Time"
   TextField "Text field_3" at 560,360 size 18x23; Text 'г.'
   TextField "Text field_4" at 337,328 size 217x23; Text 'Настройка времени ПЛК:'
   DateTimeField "Date/time field_5" at 448,395 size 111x32
      ProcessValue <- "Time_SYS_DB_SP_Time"
   DateTimeField "Date/time field_6" at 320,395 size 116x32
      ProcessValue <- "Time_SYS_DB_SP_Time"
   TextField "Text field_5" at 560,400 size 18x23; Text 'г.'
   Button "Button_1" at 320,433 size 239x32; TextOff 'Применить'
      on Click: SetBit("Time_SYS_DB_Set_Time")

screen "SIMATIC PLC system diagnostics" 800x480, template "Main"
   SysDiagControl "HmiScreenItemData" at 1,49 size 724x423
   Button "Back" at 1,1 size 159x47; TextOn 'Back'; TextOff 'Back'
      on Release: ActivateScreen("System screens", 0)

screen "System screens" 800x480, template "Main"
   Button "Back" at 1,1 size 159x47; TextOn 'Back'; TextOff 'Back'
      on Release: function_efd93a16()
   Button "HmiScreenItemData" at 36,95 size 159x47; TextOn 'SIMATIC PLC system diagnos...'; TextOff 'SIMATIC PLC system diagnos...'; PictureOn "Navigates to SIMATIC PLC system diagnostics for KTP700 Basic+ PN 14.0.1.0"; PictureOff "Navigates to SIMATIC PLC system diagnostics for KTP700 Basic+ PN 14.0.1.0"
      on Release: ActivateScreen("SIMATIC PLC system diagnostics", 0)
   Button "HmiScreenItemData_1" at 36,154 size 159x47; TextOn 'User administration'; TextOff 'User administration'; PictureOn "Navigates to User administration for KTP700 Basic+ PN 14.0.1.0"; PictureOff "Navigates to User administration for KTP700 Basic+ PN 14.0.1.0"
      on Release: ActivateScreen("User administration", 0)
   Button "HmiScreenItemData_3" at 36,272 size 159x47; TextOn 'Different jobs'; TextOff 'Different jobs'; PictureOn "Navigates to Different jobs for KTP700 Basic+ PN 14.0.1.0"; PictureOff "Navigates to Different jobs for KTP700 Basic+ PN 14.0.1.0"
      on Release: ActivateScreen("Different jobs", 0)

screen "User administration" 800x480, template "Main"
   UserView "HmiScreenItemData" at 1,49 size 724x423
   Button "Back" at 1,1 size 159x47; TextOn 'Back'; TextOff 'Back'
      on Release: ActivateScreen("System screens", 0)

Template "Settings" 800x480
   Button "Button_1" at 7,256 size 112x32; TextOff 'Привода / PolyMix_2'; Authorization "Operate"
      on Release: ActivateScreen("Dev_MD", 0); SetTag("settings", 5); SetTag("Mx", 500); SetTag("Mx_Name", 'DB 500')
      Appearance <- "settings"
   Button "Button_4" at 7,174 size 112x32; TextOff 'Сигналы - AI / Датчики'; Authorization "Operate"
      on Release: ActivateScreen("Dev_AI", 0); SetTag("settings", 3); SetTag("AIx", 300); SetTag("AIx_Name", 'DB 300')
      Appearance <- "settings"
   Button "Button_5" at 7,95 size 112x32; TextOff 'Сигналы - DI / DI'; Authorization "Operate"
      on Release: ActivateScreen("Dev_DI_1", 0); SetTag("settings", 1); SetTag("DIx", 200)
      Appearance <- "settings"
   Button "Button_27" at 7,135 size 112x32; TextOff 'Команды - DO / DO'; Authorization "Operate"
      on Release: ActivateScreen("Dev_DO_1", 0); SetTag("settings", 2); SetTag("DOx", 210)
      Appearance <- "settings"
   Button "HmiScreenItemData_1" at 7,424 size 52x47; TextOn 'System screens'; TextOff 'System'; PictureOn "Navigates to System screens for KTP700 Basic+ PN 14.0.1.0"; PictureOff "Navigates to System screens for KTP700 Basic+ PN 14.0.1.0"
      on Release: ActivateScreen("System screens", 0)
   Button "Button_3" at 7,297 size 112x32; TextOff 'Задвижки / Линии'; Authorization "Operate"
      on Release: ActivateScreen("Dev_VD2", 0); SetTag("settings", 6); SetTag("Vx", 700); SetTag("Vx_Name", 'DB 700')
      Appearance <- "settings"
   Button "Button_2" at 7,337 size 112x32; TextOff 'ШД / Задвижки'; Authorization "Operate"
      on Release: ActivateScreen("Select_Settings", 0); SetTag("settings", 7)
      Appearance <- "settings"
   Button "Button_7" at 7,216 size 112x32; TextOff 'Команды - AO / PolyMix_1'; Authorization "Operate"
      on Release: ActivateScreen("Dev_AO", 0); SetTag("settings", 4); SetTag("AOx", 400); SetTag("AOx_Name", 'DB 400')
      Appearance <- "settings"
   GraphicView "Graphic view_1" at 5,30 size 123x59; Picture "vdk3"
   TextField "Template_Text field_1" at 5,7 size 117x17; Text '+7 (495) 763-29-73'
   Button "Template_Button_1" at 4,6 size 120x84; TextOff 'Text'
      on Click: ActivateScreen("About", 0)
   Button "Button_17" at 7,376 size 112x32; TextOff 'ПИД / ШД'; Authorization "Operate"
      on Release: ActivateScreen("Dev_PID", 0); SetTag("settings", 8); SetTag("PIDx", 900); SetTag("PIDx_Name", 'DB 900')
      Appearance <- "settings"
   GraphicIOField "Template_Graphic I/O field_1" at 79,430 size 35x35; PictureList "Local_Mode"
      ProcessValue <- "Local_Mode"
   Button "Button_6" at 735,275 size 60x60; TextOff 'Text'; PictureOff "home_1"; PictureList "Alarm"
      on Click: ActivateScreen("Alarms", 0); SetTag("MainScr", 4); SetTag("Support_DB_DTR_Clean", 0)
      Appearance <- "MainScr"
      ProcessValue <- "Alm_Any"
   Button "Button_8" at 735,410 size 60x60; TextOff 'Text'; PictureOff "reset"
      on Click: SetBit("Reset_All")
   Button "Button_9" at 735,5 size 60x60; TextOff 'Text'; PictureOff "home_3"
      on Click: ActivateScreen("Root screen", 0); SetTag("MainScr", 0); SetTag("Support_DB_DTR_Clean", 0)
   Button "Button_10" at 735,5 size 60x60; TextOff 'Text'; PictureOff "home_pressed_1"
      on Click: ActivateScreen("Root screen", 0); SetTag("MainScr", 0)
      Visibility <- "MainScr"
   Button "Button_11" at 735,72 size 60x60; TextOff 'Text'; PictureOff "sett"
      on Click: SetTag("MainScr", 1); ActivateScreen("Select_Settings", 0); SetTag("settings", 0); SetTag("Support_DB_DTR_Clean", 0)
   Button "Button_12" at 735,72 size 60x60; TextOff 'Text'; PictureOff "sett_pressed"
      on Click: SetTag("MainScr", 1); ActivateScreen("Select_Settings", 0); SetTag("settings", 0); SetTag("Support_DB_DTR_Clean", 0)
      Visibility <- "MainScr"
   Button "Button_13" at 735,140 size 60x60; TextOff 'Text'; PictureOff "table"
      on Click: SetTag("MainScr", 2); ActivateScreen("Select_Alarms", 0); SetTag("Support_DB_DTR_Clean", 0)
   Button "Button_14" at 735,207 size 60x60; TextOff 'Text'; PictureOff "history"
      on Click: ActivateScreen("Select_History", 0); SetTag("MainScr", 3); SetTag("Support_DB_DTR_Clean", 0)
   Button "Button_15" at 735,140 size 60x60; TextOff 'Text'; PictureOff "table_pressed"
      on Click: SetTag("MainScr", 2); ActivateScreen("Select_Alarms", 0); SetTag("Support_DB_DTR_Clean", 0)
      Visibility <- "MainScr"
   Button "Button_16" at 735,207 size 60x60; TextOff 'Text'; PictureOff "history_pressed"
      on Click: ActivateScreen("Select_History", 0); SetTag("MainScr", 3); SetTag("Support_DB_DTR_Clean", 0)
      Appearance <- "MainScr"
      Visibility <- "MainScr"
   Button "Template_Button_2" at 735,342 size 60x60; TextOff 'Text'; PictureOff "vdk1"
      on Click: ActivateScreen("About", 0); SetTag("Support_DB_DTR_Clean", 0)

